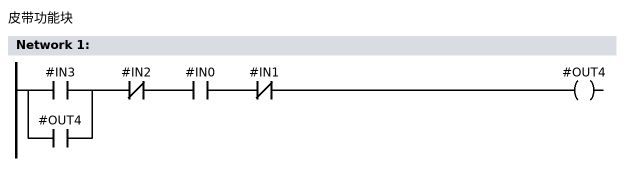
   RUNG wire#powerrail
      Contact( #IN3 )
      wire#w1
      I_Contact( #IN2 )
      Contact( #IN0 )
      I_Contact( #IN1 )
      Coil( #OUT4 )
   END_RUNG
   RUNG wire#powerrail
      Contact( #OUT4 )
   END_RUNG wire#w1
   // the same network as SCL:
   #OUT4 := (#IN3 OR #OUT4) AND NOT #IN2 AND #IN0 AND NOT #IN1;
END_REGION
END_FUNCTION

FUNCTION "脉冲累计功能块" : Void   // FC116, LAD
{ S7_Optimized_Access := 'FALSE' }
VERSION : 0.1
   VAR_INPUT
      IN0 : Bool;
      IN1 : Bool;
   END_VAR
   VAR_OUTPUT
      OUT2 : Real;
   END_VAR
   VAR_TEMP
      TEMP3 : Bool;
      TEMP4 : Real;
      TEMP5 : Real;
      TEMP6 : Real;
   END_VAR
   VAR_TEMP   // added for the SCL form of the ladder/FBD networks
      _w1 : Bool;
   END_VAR
BEGIN

REGION Network 2
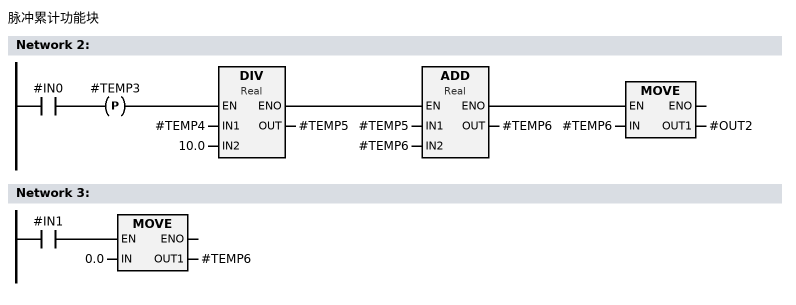
   RUNG wire#powerrail
      Contact( #IN0 )
      P_Trig( #TEMP3 )
      { S7_Templates := "SrcType := Real"; S7_GenerateENO := "TRUE" } Div(in1 := #TEMP4, in2 := 10.0, out => #TEMP5)
      { S7_Templates := "SrcType := Real"; S7_GenerateENO := "TRUE" } Add(in1 := #TEMP5, in2 := #TEMP6, out => #TEMP6)
      { S7_GenerateENO := "TRUE" } Move(in := #TEMP6, out1 => #OUT2)
   END_RUNG
   // the same network as SCL:
   // ENO of a box is taken as its EN; it also drops when the box reports an error
   #_w1 := #IN0 AND NOT #TEMP3;   // rising edge
   #TEMP3 := #IN0;
   IF #_w1 THEN
       #TEMP5 := #TEMP4 / 10.0;
       #TEMP6 := #TEMP5 + #TEMP6;
       #OUT2 := #TEMP6;
   END_IF;
END_REGION

REGION Network 3
   RUNG wire#powerrail
      Contact( #IN1 )
      { S7_GenerateENO := "TRUE" } Move(in := 0.0, out1 => #TEMP6)
   END_RUNG
   // the same network as SCL:
   IF #IN1 THEN #TEMP6 := 0.0; END_IF;
END_REGION

REGION Network 4 (STL)
         SET;
         SAVE;
END_REGION
END_FUNCTION

ORGANIZATION_BLOCK "Main"   // OB1, LAD, ProgramCycle
{ S7_Optimized_Access := 'FALSE' }
VERSION : 0.1
   VAR_TEMP
      TEMP0 : Byte;
      TEMP1 : Byte;
      TEMP2 : Byte;
      TEMP3 : Byte;
      TEMP4 : Byte;
      TEMP5 : Byte;
      TEMP6 : Int;
      TEMP7 : Int;
      TEMP8 : Int;
      TEMP9 : Date_And_Time;
   END_VAR
BEGIN

REGION Network 1
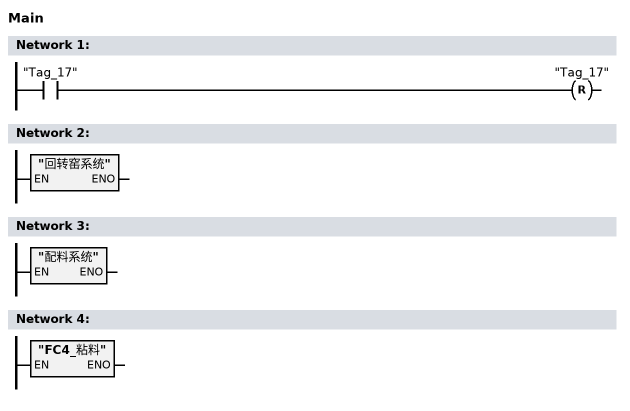
   RUNG wire#powerrail
      Contact( "Tag_17" )
      R_Coil( "Tag_17" )
   END_RUNG
   // the same network as SCL:
   IF "Tag_17" THEN "Tag_17" := FALSE; END_IF;
END_REGION

REGION Network 2
   RUNG wire#powerrail
      "回转窑系统"()
   END_RUNG
   // the same network as SCL:
   "回转窑系统"();
END_REGION

REGION Network 3
   RUNG wire#powerrail
      "配料系统"()
   END_RUNG
   // the same network as SCL:
   "配料系统"();
END_REGION

REGION Network 4
   RUNG wire#powerrail
      "FC4_粘料"()
   END_RUNG
   // the same network as SCL:
   "FC4_粘料"();
END_REGION
END_ORGANIZATION_BLOCK

ORGANIZATION_BLOCK "Cyclic interrupt"   // OB30, LAD, CyclicInterrupt
{ S7_Optimized_Access := 'TRUE' }
VERSION : 0.1
   VAR_INPUT
      Initial_Call : Bool;   // Initial call of this OB
      Event_Count : Int;   // Events discarded
   END_VAR
   VAR_TEMP   // added for the SCL form of the ladder/FBD networks
      _w1 : Bool;
      _w2 : Bool;
   END_VAR
BEGIN

REGION Network 1
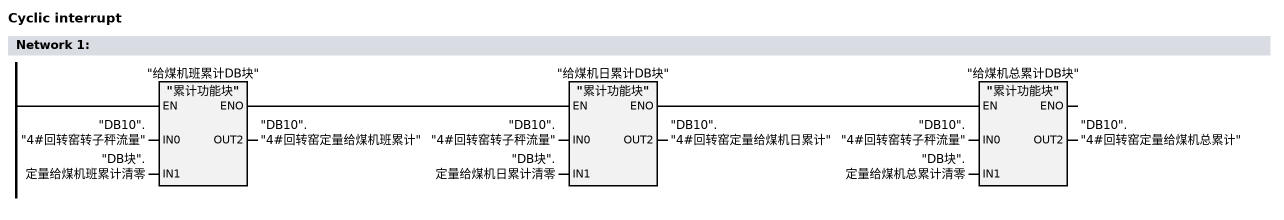
   RUNG wire#powerrail
      "给煤机班累计DB块"(IN0 := "DB10"."4#回转窑转子秤流量", IN1 := "DB块".定量给煤机班累计清零, OUT2 => "DB10"."4#回转窑定量给煤机班累计")
      "给煤机日累计DB块"(IN0 := "DB10"."4#回转窑转子秤流量", IN1 := "DB块".定量给煤机日累计清零, OUT2 => "DB10"."4#回转窑定量给煤机日累计")
      "给煤机总累计DB块"(IN0 := "DB10"."4#回转窑转子秤流量", IN1 := "DB块".定量给煤机总累计清零, OUT2 => "DB10"."4#回转窑定量给煤机总累计")
   END_RUNG
   // the same network as SCL:
   "给煤机班累计DB块"(IN0 := "DB10"."4#回转窑转子秤流量", IN1 := "DB块".定量给煤机班累计清零, OUT2 => "DB10"."4#回转窑定量给煤机班累计", ENO => #_w1);   // "累计功能块"
   "给煤机日累计DB块"(EN := #_w1,   // "累计功能块"
               IN0 := "DB10"."4#回转窑转子秤流量",
               IN1 := "DB块".定量给煤机日累计清零,
               OUT2 => "DB10"."4#回转窑定量给煤机日累计",
               ENO => #_w2);
   IF #_w2 THEN
       "给煤机总累计DB块"(IN0 := "DB10"."4#回转窑转子秤流量", IN1 := "DB块".定量给煤机总累计清零, OUT2 => "DB10"."4#回转窑定量给煤机总累计");   // "累计功能块"
   END_IF;
END_REGION
END_ORGANIZATION_BLOCK

// ===== PLC "1#LM"  CPU 1511-1 PN =====

VAR_GLOBAL   // PLC tag table "默认变量表"
   "送煤皮带备妥" AT %I0.0 : Bool;
   "送煤皮带运行" AT %I0.1 : Bool;
   "送煤皮带故障" AT %I0.2 : Bool;
   "除铁器备妥" AT %I0.3 : Bool;
   "除铁器运行" AT %I0.4 : Bool;
   "除铁器故障" AT %I0.5 : Bool;
   "定量给煤机备妥" AT %I0.6 : Bool;
   "定量给煤机运行" AT %I0.7 : Bool;
   "定量给煤机故障" AT %I1.0 : Bool;
   "煤粉收尘器备妥" AT %I1.1 : Bool;
   "煤粉收尘器运行" AT %I1.2 : Bool;
   "煤粉收尘器故障" AT %I1.3 : Bool;
   "立磨尾排风机远程" AT %I1.4 : Bool;
   "立磨尾排风机运行" AT %I1.5 : Bool;
   "立磨尾排风机故障" AT %I1.6 : Bool;
   "立磨尾排风机待机" AT %I1.7 : Bool;
   "立磨尾排高压柜远程" AT %I2.0 : Bool;
   "立磨尾排高压柜合闸" AT %I2.1 : Bool;
   "立磨尾排高压柜分闸" AT %I2.2 : Bool;
   "定量给煤机断料信号" AT %I2.3 : Bool;
   "定量给煤机左跑偏信号" AT %I2.4 : Bool;
   "定量给煤机右跑偏信号" AT %I2.5 : Bool;
   "给煤机断链信号" AT %I2.6 : Bool;
   "立磨给煤机累计脉冲" AT %I2.7 : Bool;
   "定量给料机远程" AT %I3.0 : Bool;
   "1#铰刀运行" AT %I3.1 : Bool;
   "2#铰刀运行" AT %I3.2 : Bool;
   "1#分割轮运行" AT %I3.3 : Bool;
   "2#分割轮运行" AT %I3.4 : Bool;
   "3#分割轮运行" AT %I3.5 : Bool;
   "4#分割轮运行" AT %I3.6 : Bool;
   "5#分割轮运行" AT %I3.7 : Bool;
   "立磨主机高压柜远程" AT %I4.0 : Bool;
   "立磨主机高压柜合闸" AT %I4.1 : Bool;
   "立磨主机高压柜分闸" AT %I4.2 : Bool;
   "立磨主机运行" AT %I4.3 : Bool;
   "立磨主机故障" AT %I4.4 : Bool;
   "允许主机启动" AT %I4.5 : Bool;
   "停主机" AT %I4.6 : Bool;
   "6#分割轮运行" AT %I5.0 : Bool;
   "7#分割轮运行" AT %I5.1 : Bool;
   "8#分割轮运行" AT %I5.2 : Bool;
   "9#分割轮运行" AT %I5.3 : Bool;
   "10#分割轮运行" AT %I5.4 : Bool;
   "1#灰管压力" AT %IW112 : Word;
   "2#灰管压力" AT %IW114 : Word;
   "Tag_76" AT %IW116 : Word;
   "Tag_78" AT %IW118 : Word;
   "1#母管压力USELESS" AT %IW212 : Word;
   "1#灰管压力UEELESS" AT %IW214 : Word;
   "2#母管压力USELESS" AT %IW216 : Word;
   "2#灰管压力USELESS" AT %IW218 : Word;
   "立磨尾排风机水平震动1" AT %IW256 : Int;
   "立磨尾排风机水平震动2" AT %IW258 : Int;
   "立磨尾排风机垂直震动1" AT %IW260 : Int;
   "立磨尾排风机垂直震动2" AT %IW262 : Int;
   "立磨尾排风机入口压力1" AT %IW264 : Int;
   "立磨尾排风机入口压力2" AT %IW266 : Int;
   "立磨尾排风机出口压力1" AT %IW268 : Int;
   "尾排风机入口执行器反馈" AT %IW270 : Int;
   "立磨1#煤粉仓负压" AT %IW272 : Int;
   "立磨2#煤粉仓负压" AT %IW274 : Int;
   "立磨热风管道负压" AT %IW276 : Int;
   "立磨主电机运行电流" AT %IW278 : Int;
   "立磨给煤机流量" AT %IW280 : Int;
   "立磨出口压力1" AT %IW282 : Int;
   "立磨出口压力2" AT %IW284 : Int;
   "立磨尾排风机运行转速" AT %IW288 : Int;
   "立磨尾排风机运行电流" AT %IW290 : Int;
   "立磨尾排风机出口温度1" AT %IW292 : Int;
   "立磨尾排风机入口温度1" AT %IW296 : Int;
   "立磨尾排风机入口温度2" AT %IW298 : Int;
   "立磨入磨口温度" AT %IW300 : Int;
   "1#煤粉仓1#温度" AT %ID304 : DWord;
   "1#煤粉仓2#温度" AT %ID308 : DWord;
   "1#煤粉仓3#温度" AT %ID312 : DWord;
   "1#煤粉仓4#温度" AT %ID316 : DWord;
   "1#煤粉仓5#温度" AT %ID320 : DWord;
   "1#煤粉仓6#温度" AT %ID324 : DWord;
   "2#煤粉仓1#温度" AT %ID328 : DWord;
   "2#煤粉仓2#温度" AT %ID332 : DWord;
   "2#煤粉仓3#温度" AT %ID336 : DWord;
   "2#煤粉仓4#温度" AT %ID340 : DWord;
   "2#煤粉仓5#温度" AT %ID344 : DWord;
   "2#煤粉仓6#温度" AT %ID348 : DWord;
   "电机绕组U相温度" AT %ID352 : DWord;
   "电机绕组V相温度" AT %ID356 : DWord;
   "电机绕组W相温度" AT %ID360 : DWord;
   "尾排电机前轴温度" AT %ID364 : DWord;
   "尾排电机后轴温度" AT %ID368 : DWord;
   "尾排风机前轴温度" AT %ID372 : DWord;
   "尾排风机后轴温度" AT %ID376 : DWord;
   "立磨机出口温度1" AT %ID380 : DWord;
   "立磨机出口温度2" AT %ID384 : DWord;
   "Tag_101" AT %ID388 : DWord;
   "Tag_102" AT %ID392 : DWord;
   "Tag_103" AT %ID396 : DWord;
   "送煤皮带驱动" AT %Q0.0 : Bool;
   "除铁器驱动" AT %Q0.1 : Bool;
   "定量给煤机驱动" AT %Q0.2 : Bool;
   "煤粉收尘器驱动" AT %Q0.3 : Bool;
   "立磨尾排风机停止" AT %Q0.4 : Bool;
   "立磨尾排高压柜合闸驱动" AT %Q0.5 : Bool;
   "立磨尾排风机高压柜分闸" AT %Q0.6 : Bool;
   "立磨尾排风机驱动" AT %Q0.7 : Bool;
   "立磨主机高压柜合闸驱动" AT %Q1.0 : Bool;
   "立磨主机高压柜分闸驱动" AT %Q1.1 : Bool;
   "Tag_107" AT %QB4 : Byte;
   "1#仓泵手/自动" AT %Q100.0 : Bool;
   "1#仓泵自动启动" AT %Q100.1 : Bool;
   "1#仓泵自动停止" AT %Q100.2 : Bool;
   "2#仓泵手/自动" AT %Q100.3 : Bool;
   "2#仓泵自动启动" AT %Q100.4 : Bool;
   "2#仓泵自动停止" AT %Q100.5 : Bool;
   "1#排气阀手动开" AT %Q101.0 : Bool;
   "1#排气阀手动关" AT %Q101.1 : Bool;
   "1#进料阀手动开" AT %Q101.2 : Bool;
   "1#进料阀手动关" AT %Q101.3 : Bool;
   "1#出料阀手动开" AT %Q101.4 : Bool;
   "1#出料阀手动关" AT %Q101.5 : Bool;
   "1#进气阀手动开" AT %Q101.6 : Bool;
   "1#进气阀手动关" AT %Q101.7 : Bool;
   "1#助吹阀手动开" AT %Q102.0 : Bool;
   "1#助吹阀手动关" AT %Q102.1 : Bool;
   "1#排堵阀手动开" AT %Q102.2 : Bool;
   "1#排堵阀手动关" AT %Q102.3 : Bool;
   "2#排气阀手动开" AT %Q102.4 : Bool;
   "2#排气阀手动关" AT %Q102.5 : Bool;
   "2#进料阀手动开" AT %Q102.6 : Bool;
   "2#进料阀手动关" AT %Q102.7 : Bool;
   "2#出料阀手动开" AT %Q103.0 : Bool;
   "2#出料阀手动关" AT %Q103.1 : Bool;
   "2#进气阀手动开" AT %Q103.2 : Bool;
   "2#进气阀手动关" AT %Q103.3 : Bool;
   "2#助吹阀手动开" AT %Q103.4 : Bool;
   "2#助吹阀手动关" AT %Q103.5 : Bool;
   "2#排堵阀手动开" AT %Q103.6 : Bool;
   "2#排堵阀手动关" AT %Q103.7 : Bool;
   "1#切1#切换阀手动开" AT %Q104.0 : Bool;
   "1#切1#切换阀手动关" AT %Q104.1 : Bool;
   "1#切2#切换阀手动开" AT %Q104.2 : Bool;
   "1#切2#切换阀手动关" AT %Q104.3 : Bool;
   "1#切3#切换阀手动开" AT %Q104.4 : Bool;
   "1#切3#切换阀手动关" AT %Q104.5 : Bool;
   "1#切4#切换阀手动开" AT %Q104.6 : Bool;
   "1#切4#切换阀手动关" AT %Q104.7 : Bool;
   "1#切5#切换阀手动开" AT %Q105.0 : Bool;
   "1#切5#切换阀手动关" AT %Q105.1 : Bool;
   "2#切1#切换阀手动开" AT %Q105.2 : Bool;
   "2#切1#切换阀手动关" AT %Q105.3 : Bool;
   "2#切2#切换阀手动开" AT %Q105.4 : Bool;
   "1#母管压力下限" AT %QW108 : Word;
   "1#灰管压力下限" AT %QW110 : Word;
   "1#灰管压力上限" AT %QW112 : Word;
   "1#进料时间" AT %QW114 : Word;
   "1#吹扫时间" AT %QW116 : Word;
   "2#母管压力下限" AT %QW118 : Word;
   "2#灰管压力下限" AT %QW120 : Word;
   "2#灰管压力上限" AT %QW122 : Word;
   "2#进料时间" AT %QW124 : Word;
   "立磨给煤机流量给定" AT %QW256 : Int;
   "立磨尾排风机转速给定" AT %QW258 : Int;
   "尾排风机入口执行器给定" AT %QW260 : Int;
   "Tag_5" AT %M2.0 : Bool;
   "Tag_11" AT %M2.3 : Bool;
   "Tag_19" AT %M2.5 : Bool;
   "Tag_1" AT %MW4 : Word;
   "Tag_8" AT %MW10 : Word;
   "Tag_6" AT %MW12 : Word;
   "Tag_21" AT %MW14 : Word;
   "Tag_16" AT %MW16 : Word;
   "锁风定量给煤机流量累计清零" AT %M30.1 : Bool;
   "Tag_13" AT %MW100 : Word;
   "Tag_12" AT %M300.0 : Bool;
   "Tag_20" AT %M300.1 : Bool;
   "Tag_9" AT %M400.0 : Bool;
   "Tag_17" AT %M400.1 : Bool;
   "1#仓泵进料时间" AT %MW506 : Word;
   "1#仓泵吹扫时间" AT %MW508 : Word;
   "1#母管下限" AT %MW510 : Word;
   "1#灰管上限" AT %MW512 : Word;
   "1#灰管下限" AT %MW514 : Word;
   "2#仓泵进料时间" AT %MW516 : Word;
   "2#仓泵吹扫时间" AT %MW518 : Word;
   "2#母管下限" AT %MW520 : Word;
   "2#灰管上限" AT %MW522 : Word;
   "2#灰管下限" AT %MW524 : Word;
   "1#母管压力信号" AT %MW526 : Word;
   "1#灰管压力信号" AT %MW528 : Word;
   "2#母管压力信号" AT %MW530 : Word;
   "2#灰管压力信号" AT %MW532 : Word;
   "1#仓泵手自动标示" AT %M600.1 : Bool;
   "2#仓泵手自动标示" AT %M600.2 : Bool;
   "Tag_3" AT %T100 : Timer;
   "Tag_4" AT %T101 : Timer;
   "Tag_10" AT %C1 : Counter;
   "Tag_18" AT %C2 : Counter;
   "I4_7" AT %I4.7 : Bool;
   "I5_5" AT %I5.5 : Bool;
   "I5_6" AT %I5.6 : Bool;
   "I5_7" AT %I5.7 : Bool;
   "1#板式给煤机-褐煤备妥" AT %I6.0 : Bool;
   "1#板式给煤机-褐煤运行" AT %I6.1 : Bool;
   "1#板式给煤机-褐煤故障" AT %I6.2 : Bool;
   "2#板式给煤机-烟煤备妥" AT %I6.3 : Bool;
   "2#板式给煤机-烟煤运行" AT %I6.4 : Bool;
   "2#板式给煤机-烟煤故障" AT %I6.5 : Bool;
   "I6_6" AT %I6.6 : Bool;
   "I6_7" AT %I6.7 : Bool;
   "I7_0" AT %I7.0 : Bool;
   "I7_1" AT %I7.1 : Bool;
   "I7_2" AT %I7.2 : Bool;
   "I7_3" AT %I7.3 : Bool;
   "I7_4" AT %I7.4 : Bool;
   "I7_5" AT %I7.5 : Bool;
   "I7_6" AT %I7.6 : Bool;
   "I7_7" AT %I7.7 : Bool;
   "I8_0" AT %I8.0 : Bool;
   "I8_1" AT %I8.1 : Bool;
   "I8_2" AT %I8.2 : Bool;
   "I8_3" AT %I8.3 : Bool;
   "I8_4" AT %I8.4 : Bool;
   "I8_5" AT %I8.5 : Bool;
   "I8_6" AT %I8.6 : Bool;
   "I8_7" AT %I8.7 : Bool;
   "I9_0" AT %I9.0 : Bool;
   "I9_1" AT %I9.1 : Bool;
   "I9_2" AT %I9.2 : Bool;
   "I9_3" AT %I9.3 : Bool;
   "I9_4" AT %I9.4 : Bool;
   "I9_5" AT %I9.5 : Bool;
   "I9_6" AT %I9.6 : Bool;
   "I9_7" AT %I9.7 : Bool;
   "I10_0" AT %I10.0 : Bool;
   "I10_1" AT %I10.1 : Bool;
   "I10_2" AT %I10.2 : Bool;
   "I10_3" AT %I10.3 : Bool;
   "I10_4" AT %I10.4 : Bool;
   "I10_5" AT %I10.5 : Bool;
   "I10_6" AT %I10.6 : Bool;
   "I10_7" AT %I10.7 : Bool;
   "I11_0" AT %I11.0 : Bool;
   "I11_1" AT %I11.1 : Bool;
   "I11_2" AT %I11.2 : Bool;
   "I11_3" AT %I11.3 : Bool;
   "I11_4" AT %I11.4 : Bool;
   "I11_5" AT %I11.5 : Bool;
   "I11_6" AT %I11.6 : Bool;
   "I11_7" AT %I11.7 : Bool;
   "1#板式给煤机-褐煤启停" AT %Q1.2 : Bool;
   "2#板式给煤机-烟煤启停" AT %Q1.3 : Bool;
   "立磨现场皮带报警器" AT %Q1.4 : Bool;
   "立磨中控报警器" AT %Q1.5 : Bool;
   "Q1_6" AT %Q1.6 : Bool;
   "Q1_7" AT %Q1.7 : Bool;
   "Q2_0" AT %Q2.0 : Bool;
   "Q2_1" AT %Q2.1 : Bool;
   "Q2_2" AT %Q2.2 : Bool;
   "Q2_3" AT %Q2.3 : Bool;
   "Q2_4" AT %Q2.4 : Bool;
   "Q2_5" AT %Q2.5 : Bool;
   "Q2_6" AT %Q2.6 : Bool;
   "Q2_7" AT %Q2.7 : Bool;
   "Q3_0" AT %Q3.0 : Bool;
   "Q3_1" AT %Q3.1 : Bool;
   "Q3_2" AT %Q3.2 : Bool;
   "Q3_3" AT %Q3.3 : Bool;
   "Q3_4" AT %Q3.4 : Bool;
   "Q3_5" AT %Q3.5 : Bool;
   "Q3_6" AT %Q3.6 : Bool;
   "Q3_7" AT %Q3.7 : Bool;
   "1#板式给煤机-褐煤流量反馈" AT %IW286 : Int;
   "2#板式给煤机-烟煤流量反馈" AT %IW294 : Int;
   "PIW302" AT %IW302 : Int;
   "1#板式给煤机-褐煤流量给定" AT %QW262 : Int;
   "2#板式给煤机-烟煤流量给定" AT %QW264 : Int;
   "PQW266" AT %QW266 : Int;
   "PQW268" AT %QW268 : Int;
   "PQW270" AT %QW270 : Int;
   "立磨煤粉仓称重" AT %ID400 : Real;
   "立磨1#煤粉仓称重" AT %ID408 : Real;
   "立磨2#煤粉仓称重" AT %ID416 : Real;
   "1#立磨板式给料流量累计清零" AT %M30.2 : Bool;
   "2#立磨板式给料流量累计清零" AT %M30.3 : Bool;
   "Tag_2" AT %M30.7 : Bool;
   "Tag_80" AT %M80.0 : Bool;
   "Tag_81" AT %M81.0 : Bool;
   "Tag_82" AT %M80.1 : Bool;
   "Tag_83" AT %M80.2 : Bool;
   "Tag_84" AT %M80.3 : Bool;
   "Tag_85" AT %M81.1 : Bool;
   "Tag_86" AT %T102 : Timer;
   "Clock_Byte" AT %MB0 : Byte;
   "Clock_10Hz" AT %M0.0 : Bool;
   "Clock_5Hz" AT %M0.1 : Bool;
   "Clock_2.5Hz" AT %M0.2 : Bool;
   "Clock_2Hz" AT %M0.3 : Bool;
   "Clock_1.25Hz" AT %M0.4 : Bool;
   "Clock_1Hz" AT %M0.5 : Bool;
   "Clock_0.625Hz" AT %M0.6 : Bool;
   "Clock_0.5Hz" AT %M0.7 : Bool;
   "System_Byte" AT %MB1 : Byte;
   "FirstScan" AT %M1.0 : Bool;
   "DiagStatusUpdate" AT %M1.1 : Bool;
   "AlwaysTRUE" AT %M1.2 : Bool;
   "AlwaysFALSE" AT %M1.3 : Bool;
   "2#切2#切换阀手动关" AT %Q105.5 : Bool;
   "3#切1#切换阀手动开" AT %Q105.6 : Bool;
   "3#切1#切换阀手动关" AT %Q105.7 : Bool;
   "3#切2#切换阀手动开" AT %Q106.0 : Bool;
   "3#切2#切换阀手动关" AT %Q106.1 : Bool;
   "4#切1#切换阀手动开" AT %Q106.2 : Bool;
   "4#切1#切换阀手动关" AT %Q106.3 : Bool;
   "4#切2#切换阀手动开" AT %Q106.4 : Bool;
   "4#切2#切换阀手动关" AT %Q106.5 : Bool;
   "4#切3#切换阀手动开" AT %Q106.6 : Bool;
   "4#切3#切换阀手动关" AT %Q106.7 : Bool;
   "4#切4#切换阀手动开" AT %Q107.0 : Bool;
   "4#切4#切换阀手动关" AT %Q107.1 : Bool;
   "Tag_20(1)" AT %Q107.2 : Bool;
   "Tag_21(1)" AT %Q107.3 : Bool;
   "Tag_22" AT %Q107.4 : Bool;
   "Tag_23" AT %Q107.5 : Bool;
   "Tag_24" AT %Q107.6 : Bool;
   "Tag_25" AT %Q107.7 : Bool;
   "2#吹扫时间" AT %QW126 : Word;
   "1#排气阀关到位" AT %I100.0 : Bool;
   "1#排气阀开到位" AT %I100.1 : Bool;
   "1#进料阀关到位" AT %I100.2 : Bool;
   "1#进料阀开到位" AT %I100.3 : Bool;
   "1#出料阀关到位" AT %I100.4 : Bool;
   "1#出料阀开到位" AT %I100.5 : Bool;
   "1#进气阀关到位" AT %I100.6 : Bool;
   "1#进气阀开到位" AT %I100.7 : Bool;
   "1#助吹阀关到位" AT %I101.0 : Bool;
   "1#助吹阀开到位" AT %I101.1 : Bool;
   "1#排堵阀关到位" AT %I101.2 : Bool;
   "1#排堵阀开到位" AT %I101.3 : Bool;
   "1#料位信号" AT %I101.4 : Bool;
   "1#现场箱远程" AT %I101.5 : Bool;
   "2#排气阀关到位" AT %I101.6 : Bool;
   "2#排气阀开到位" AT %I101.7 : Bool;
   "2#进料阀关到位" AT %I102.0 : Bool;
   "2#进料阀开到位" AT %I102.1 : Bool;
   "2#出料阀关到位" AT %I102.2 : Bool;
   "2#出料阀开到位" AT %I102.3 : Bool;
   "2#进气阀关到位" AT %I102.4 : Bool;
   "2#进气阀开到位" AT %I102.5 : Bool;
   "2#助吹阀关到位" AT %I102.6 : Bool;
   "2#助吹阀开到位" AT %I102.7 : Bool;
   "2#排堵阀关到位" AT %I103.0 : Bool;
   "2#排堵阀开到位" AT %I103.1 : Bool;
   "2#料位信号" AT %I103.2 : Bool;
   "2#现场箱远程" AT %I103.3 : Bool;
   "1#切1#切换阀关到位" AT %I103.4 : Bool;
   "1#切1#切换阀开到位" AT %I103.5 : Bool;
   "1#切2#切换阀关到位" AT %I103.6 : Bool;
   "1#切2#切换阀开到位" AT %I103.7 : Bool;
   "1#切3#切换阀关到位" AT %I104.0 : Bool;
   "1#切3#切换阀开到位" AT %I104.1 : Bool;
   "1#切4#切换阀关到位" AT %I104.2 : Bool;
   "1#切4#切换阀开到位" AT %I104.3 : Bool;
   "1#切5#切换阀关到位" AT %I104.4 : Bool;
   "1#切5#切换阀开到位" AT %I104.5 : Bool;
   "1#切远程信号" AT %I104.6 : Bool;
   "2#切1#切换阀关到位" AT %I104.7 : Bool;
   "2#切1#切换阀开到位" AT %I105.0 : Bool;
   "2#切2#切换阀关到位" AT %I105.1 : Bool;
   "2#切2#切换阀开到位" AT %I105.2 : Bool;
   "2#切远程信号" AT %I105.3 : Bool;
   "3#切1#切换阀关到位" AT %I105.4 : Bool;
   "3#切1#切换阀开到位" AT %I105.5 : Bool;
   "3#切2#切换阀关到位" AT %I105.6 : Bool;
   "3#切2#切换阀开到位" AT %I105.7 : Bool;
   "3#切远程信号" AT %I106.0 : Bool;
   "4#切1#切换阀关到位" AT %I106.1 : Bool;
   "4#切1#切换阀开到位" AT %I106.2 : Bool;
   "4#切2#切换阀关到位" AT %I106.3 : Bool;
   "4#切2#切换阀开到位" AT %I106.4 : Bool;
   "4#切3#切换阀关到位" AT %I106.5 : Bool;
   "4#切3#切换阀开到位" AT %I106.6 : Bool;
   "4#切4#切换阀关到位" AT %I106.7 : Bool;
   "4#切4#切换阀开到位" AT %I107.0 : Bool;
   "4#切远程信号" AT %I107.1 : Bool;
   "1#中控备妥" AT %I107.2 : Bool;
   "1#运行" AT %I107.3 : Bool;
   "1#母管压力低" AT %I107.4 : Bool;
   "1#灰管压力高" AT %I107.5 : Bool;
   "2#中控备妥" AT %I107.6 : Bool;
   "2#运行" AT %I107.7 : Bool;
   "2#母管压力低" AT %I108.0 : Bool;
   "2#灰管压力高" AT %I108.1 : Bool;
   "Tag_7" AT %MW200 : Word;
   "Tag_14" AT %MW202 : Word;
   "Tag_15" AT %M200.0 : Bool;
   "Tag_26" AT %M200.1 : Bool;
   "Tag_27" AT %Q4.0 : Bool;
   "Tag_28" AT %M2.1 : Bool;
   "Tag_29" AT %MW82 : Word;
   "Tag_30" AT %C3 : Counter;
   "Tag_31" AT %C4 : Counter;
   "母管压力" AT %IW110 : Word;
   "Tag_32" AT %M10.0 : Bool;
   "Tag_33" AT %MD40 : Real;
   "Tag_34" AT %MD44 : Real;
   "Tag_35" AT %MD48 : Real;
   "Tag_36" AT %M60.0 : Bool;
   "HMI_ALARM_RST" AT %M10.1 : Bool;
   "Tag_38" AT %M10.2 : Bool;
END_VAR

DATA_BLOCK "qud"   // DB1
{ S7_Optimized_Access := 'FALSE' }
VERSION : 0.1
   VAR
      STAT0 : Bool;
      STAT1 : Bool;
      STAT2 : Bool;
      STAT3 : Bool;
      STAT4 : Bool;
      STAT5 : Bool;
      STAT6 : Bool;
      STAT7 : Bool;
      STAT8 : Bool;
      STAT9 : Bool;
      STAT10 : Bool;
      STAT11 : Bool;
      STAT12 : Bool;
      STAT13 : Bool;
      STAT14 : Bool;
      STAT15 : Bool;
      "1#立磨板式给料机启动" : Bool;
      "1#立磨板式给料机停止" : Bool;
      "2#立磨板式给料机启动" : Bool;
      "2#立磨板式给料机停止" : Bool;
      STAT20 : Bool;
      STAT21 : Bool;
      STAT22 : Bool;
      STAT23 : Bool;
   END_VAR
BEGIN
END_DATA_BLOCK

DATA_BLOCK "MNL"   // DB2
{ S7_Optimized_Access := 'FALSE' }
VERSION : 0.1
   VAR
      锁风定量给煤机 : Real := 44.0;
      锁风定量给煤机流量反馈 : Real;
      立磨尾排水平振动1 : Real;
      立磨尾排水平振动2 : Real;
      立磨尾排风机垂直振动1 : Real;
      立磨尾排风机垂直振动2 : Real;
      立磨尾排风机出口压力1 : Real;
      立磨尾排风机出口压力2 : Real;
      STAT8 : Real := 56.07639;
      立磨尾排风机出口温度2 : Real;
      STAT10 : Real := 47.39583;
      STAT11 : Real := 46.52778;
      立磨尾排风机入口压力1 : Real := -2147.512;
      立磨尾排风机入口压力2 : Real := -2461.689;
      "立磨1#煤粉仓负压" : Real := -300.0;
      "立磨2#煤粉仓负压" : Real := -272.9167;
      立磨热风管道负压 : Real := -562.5;
      立磨煤粉仓称重 : Real := 101.51;
      "立磨1#煤粉仓称重" : Real := 8.44;
      "立磨2#煤粉仓称重" : Real := 13.24;
      尾排风机运行频率 : Real := 744.2824;
      尾排风机运行电流 : Real := 41.25;
      主电机运行电流 : Real;
      立磨尾排风机转速给定 : Real := 500.0;
      锁风定量给煤机流量累计 : Real := 30006.97;
      "1#煤粉仓1#温度" : Real := 37.0;
      "1#煤粉仓2#温度" : Real := 36.0;
      "1#煤粉仓3#温度" : Real := 37.0;
      "1#煤粉仓4#温度" : Real := 36.0;
      "1#煤粉仓5#温度" : Real := 36.0;
      "1#煤粉仓6#温度" : Real := 37.0;
      "2#煤粉仓1#温度" : Real := 37.0;
      "2#煤粉仓2#温度" : Real := 36.0;
      "2#煤粉仓3#温度" : Real := 37.0;
      "2#煤粉仓4#温度" : Real := 37.0;
      "2#煤粉仓5#温度" : Real := 37.0;
      "2#煤粉仓6#温度" : Real := 37.0;
      电机绕组U相温度 : Real := 59.0;
      电机绕组V相温度 : Real := 57.0;
      电机绕组W相温度 : Real := 59.0;
      尾排电机前轴温度 : Real := 34.0;
      尾排电机后轴温度 : Real := 40.0;
      尾排风机前轴温度 : Real := 144.8206;
      尾排风机后轴温度 : Real;
      立磨机出口温度1 : Real;
      立磨机出口温度2 : Real := 43.0;
      STAT46 : Real := 46.0;
      STAT47 : Real := 62.0;
      STAT48 : Real := 58.0;
      立磨尾排风机出口温度1 : Real := -1753.472;
      立磨尾排风机入口温度1 : Real := -1707.176;
      立磨尾排风机入口温度2 : Real;
      尾排风机执行器开度给定 : Real;
      尾排风机执行器开度反馈 : Real;
      立磨机出口压力1 : Real;
      立磨机出口压力2 : Real;
      立磨主电机入磨口温度 : Real;
      "1#立磨板式给料反馈" : Real;
      "2#立磨板式给料反馈" : Real;
      "1#立磨板式给料给定" : Real;
      "2#立磨板式给料给定" : Real;
      "1#立磨板式给料累计" : Real;
      "2#立磨板式给料累计" : Real;
      STAT63 : Real;
      STAT64 : Real;
      STAT65 : Real;
   END_VAR
BEGIN
END_DATA_BLOCK

DATA_BLOCK "TIMEDB"   // DB3
{ S7_Optimized_Access := 'TRUE' }
VERSION : 0.1
   VAR
      T1 : IEC_TIMER;
      T2 : IEC_TIMER;
      T3 : IEC_TIMER;
      T4 : IEC_TIMER;
      T5 : IEC_TIMER;
      T6 : IEC_TIMER;
      T7 : IEC_TIMER;
      T8 : IEC_TIMER;
      T9 : IEC_TIMER;
      T10 : IEC_TIMER;
      T11 : IEC_TIMER;
      T12 : IEC_TIMER;
      T13 : IEC_TIMER;
      T14 : IEC_TIMER;
      T15 : IEC_TIMER;
      T16 : IEC_TIMER;
      T17 : IEC_TIMER;
      T18 : IEC_TIMER;
      T19 : IEC_TIMER;
      T20 : IEC_TIMER;
      T21 : IEC_TIMER;
      T22 : IEC_TIMER;
      T23 : IEC_TIMER;
      T24 : IEC_TIMER;
      T25 : IEC_TIMER;
      T26 : IEC_TIMER;
      T27 : IEC_TIMER;
      T28 : IEC_TIMER;
      T29 : IEC_TIMER;
      T30 : IEC_TIMER;
      T31 : IEC_TIMER;
      T32 : IEC_TIMER;
      T33 : IEC_TIMER;
      T34 : IEC_TIMER;
      T35 : IEC_TIMER;
      T36 : IEC_TIMER;
      T37 : IEC_TIMER;
      T38 : IEC_TIMER;
      T39 : IEC_TIMER;
      T40 : IEC_TIMER;
      T41 : IEC_TIMER;
      T42 : IEC_TIMER;
      T43 : IEC_TIMER;
      T44 : IEC_TIMER;
      T45 : IEC_TIMER;
      T46 : IEC_TIMER;
      T47 : IEC_TIMER;
      T48 : IEC_TIMER;
      T49 : IEC_TIMER;
      T50 : IEC_TIMER;
      T51 : IEC_TIMER;
      T52 : IEC_TIMER;
      T53 : IEC_TIMER;
      T54 : IEC_TIMER;
      T55 : IEC_TIMER;
      T56 : IEC_TIMER;
      T57 : IEC_TIMER;
      T58 : IEC_TIMER;
      T59 : IEC_TIMER;
      T60 : IEC_TIMER;
      T61 : IEC_TIMER;
      T62 : IEC_TIMER;
      T63 : IEC_TIMER;
      T64 : IEC_TIMER;
      T65 : IEC_TIMER;
      T66 : IEC_TIMER;
      T67 : IEC_TIMER;
      T68 : IEC_TIMER;
      T69 : IEC_TIMER;
      T70 : IEC_TIMER;
      T71 : IEC_TIMER;
      T72 : IEC_TIMER;
      T73 : IEC_TIMER;
      T74 : IEC_TIMER;
      T75 : IEC_TIMER;
      T76 : IEC_TIMER;
      T77 : IEC_TIMER;
      T78 : IEC_TIMER;
      T79 : IEC_TIMER;
      T80 : IEC_TIMER;
      T81 : IEC_TIMER;
      T82 : IEC_TIMER;
      T83 : IEC_TIMER;
      T84 : IEC_TIMER;
      T85 : IEC_TIMER;
      T86 : IEC_TIMER;
      T87 : IEC_TIMER;
      T88 : IEC_TIMER;
      T89 : IEC_TIMER;
      T90 : IEC_TIMER;
      T91 : IEC_TIMER;
      T92 : IEC_TIMER;
      T93 : IEC_TIMER;
      T94 : IEC_TIMER;
      T95 : IEC_TIMER;
      T96 : IEC_TIMER;
      T97 : IEC_TIMER;
      T98 : IEC_TIMER;
      T99 : IEC_TIMER;
      T100 : IEC_TIMER;
   END_VAR
BEGIN
END_DATA_BLOCK

DATA_BLOCK "累计功能块_DB_1"   // DB4
{ S7_Optimized_Access := 'FALSE' }
VERSION : 0.1
// stored: InstanceOfName 累计功能块
"累计功能块"
BEGIN
END_DATA_BLOCK

DATA_BLOCK "累计功能块_DB"   // DB5
{ S7_Optimized_Access := 'FALSE' }
VERSION : 0.1
// stored: InstanceOfName 累计功能块
"累计功能块"
BEGIN
END_DATA_BLOCK

DATA_BLOCK "累计功能块_DB_2"   // DB6
{ S7_Optimized_Access := 'FALSE' }
VERSION : 0.1
// stored: InstanceOfName 累计功能块
"累计功能块"
BEGIN
END_DATA_BLOCK

DATA_BLOCK "DB9_P"   // DB9
{ S7_Optimized_Access := 'FALSE' }
VERSION : 0.1
   VAR
      P1 : Bool;
      P2 : Bool;
      P3 : Bool;
      P4 : Bool;
      P5 : Bool;
      P6 : Bool;
      P7 : Bool;
      P8 : Bool;
      P9 : Bool;
      P10 : Bool;
      P11 : Bool;
      P12 : Bool;
      P13 : Bool;
      P14 : Bool;
      P15 : Bool;
      P16 : Bool;
      P17 : Bool;
      P18 : Bool;
      P19 : Bool;
      P20 : Bool;
      P21 : Bool;
      P22 : Bool;
      P23 : Bool;
      P24 : Bool;
      P25 : Bool;
      P26 : Bool;
      P27 : Bool;
      P28 : Bool;
      P29 : Bool;
      P30 : Bool;
      P31 : Bool;
      P32 : Bool;
      P33 : Bool;
      P34 : Bool;
      P35 : Bool;
      P36 : Bool;
      P37 : Bool;
      P38 : Bool;
      P39 : Bool;
      P40 : Bool;
      P41 : Bool;
      P42 : Bool;
      P43 : Bool;
      P44 : Bool;
      P45 : Bool;
      P46 : Bool;
      P47 : Bool;
      P48 : Bool;
      P49 : Bool;
      P50 : Bool;
      P51 : Bool;
      P52 : Bool;
      P53 : Bool;
      P54 : Bool;
      P55 : Bool;
      P56 : Bool;
      P57 : Bool;
      P58 : Bool;
      P59 : Bool;
      P60 : Bool;
      P61 : Bool;
      P62 : Bool;
      P63 : Bool;
      P64 : Bool;
      P65 : Bool;
      P66 : Bool;
      P67 : Bool;
      P68 : Bool;
      P69 : Bool;
      P70 : Bool;
      P71 : Bool;
      P72 : Bool;
      P73 : Bool;
      P74 : Bool;
      P75 : Bool;
      P76 : Bool;
      P77 : Bool;
      P78 : Bool;
      P79 : Bool;
      P80 : Bool;
      P81 : Bool;
      P82 : Bool;
      P83 : Bool;
      P84 : Bool;
      P85 : Bool;
      P86 : Bool;
      P87 : Bool;
      P88 : Bool;
      P89 : Bool;
      P90 : Bool;
      P91 : Bool;
      P92 : Bool;
      P93 : Bool;
   END_VAR
BEGIN
END_DATA_BLOCK

DATA_BLOCK "HMI_IN_BOOL"   // DB10
{ S7_Optimized_Access := 'FALSE' }
VERSION : 0.1
   VAR
      "1#仓泵手/自动" : Bool;
      "1#仓泵自动启动" : Bool;
      "1#仓泵自动停止" : Bool;
      "2#仓泵手/自动" : Bool;
      "2#仓泵自动启动" : Bool;
      "2#仓泵自动停止" : Bool;
      DB10_0_6 : Bool;
      DB10_0_7 : Bool;
      "1#排气阀手动开" : Bool;
      "1#排气阀手动关" : Bool;
      "1#进料阀手动开" : Bool;
      "1#进料阀手动关" : Bool;
      "1#出料阀手动开" : Bool;
      "1#出料阀手动关" : Bool;
      "1#进气阀手动开" : Bool;
      "1#进气阀手动关" : Bool;
      "1#助吹阀手动开" : Bool;
      "1#助吹阀手动关" : Bool;
      "1#排堵阀手动开" : Bool;
      "1#排堵阀手动关" : Bool;
      "2#排气阀手动开" : Bool;
      "2#排气阀手动关" : Bool;
      "2#进料阀手动开" : Bool;
      "2#进料阀手动关" : Bool;
      "2#出料阀手动开" : Bool;
      "2#出料阀手动关" : Bool;
      "2#进气阀手动开" : Bool;
      "2#进气阀手动关" : Bool;
      "2#助吹阀手动开" : Bool;
      "2#助吹阀手动关" : Bool;
      "2#排堵阀手动开" : Bool;
      "2#排堵阀手动关" : Bool;
      "1#切1#切换阀手动开" : Bool;
      "1#切1#切换阀手动关" : Bool;
      "1#切2#切换阀手动开" : Bool;
      "1#切2#切换阀手动关" : Bool;
      "1#切3#切换阀手动开" : Bool;
      "1#切3#切换阀手动关" : Bool;
      "1#切4#切换阀手动开" : Bool;
      "1#切4#切换阀手动关" : Bool;
      "1#切5#切换阀手动开" : Bool;
      "1#切5#切换阀手动关" : Bool;
      "2#切1#切换阀手动开" : Bool;
      "2#切1#切换阀手动关" : Bool;
      "2#切2#切换阀手动开" : Bool;
      "2#切2#切换阀手动关" : Bool;
      "3#切1#切换阀手动开" : Bool;
      "3#切1#切换阀手动关" : Bool;
      "3#切2#切换阀手动开" : Bool;
      "3#切2#切换阀手动关" : Bool;
      "4#切1#切换阀手动开" : Bool;
      "4#切1#切换阀手动关" : Bool;
      "4#切2#切换阀手动开" : Bool;
      "4#切2#切换阀手动关" : Bool;
      "4#切3#切换阀手动开" : Bool;
      "4#切3#切换阀手动关" : Bool;
      "4#切4#切换阀手动开" : Bool;
      "4#切4#切换阀手动关" : Bool;
      DB10_7_2 : Bool;
      DB10_7_3 : Bool;
      DB10_7_4 : Bool;
      DB10_7_5 : Bool;
      DB10_7_6 : Bool;
      DB10_7_7 : Bool;
      DB10_8_0 : Bool;
      DB10_8_1 : Bool;
      DB10_8_2 : Bool;
      DB10_8_3 : Bool;
      DB10_8_4 : Bool;
      DB10_8_5 : Bool;
      DB10_8_6 : Bool;
      DB10_8_7 : Bool;
      DB10_9_0 : Bool;
      DB10_9_1 : Bool;
      DB10_9_2 : Bool;
      DB10_9_3 : Bool;
      DB10_9_4 : Bool;
      DB10_9_5 : Bool;
      DB10_9_6 : Bool;
      DB10_9_7 : Bool;
      DB10_10_0 : Bool;
      DB10_10_1 : Bool;
      DB10_10_2 : Bool;
      DB10_10_3 : Bool;
      DB10_10_4 : Bool;
      DB10_10_5 : Bool;
      DB10_10_6 : Bool;
      DB10_10_7 : Bool;
      DB_10_11_0 : Bool;
      DB_10_11_1 : Bool;
      DB_10_11_2 : Bool;
      DB_10_11_3 : Bool;
      DB_10_11_4 : Bool;
      DB_10_11_5 : Bool;
      DB_10_11_6 : Bool;
      DB_10_11_7 : Bool;
      DB_10_11_8 : Bool;
      DB_10_11_9 : Bool;
      DB_10_11_10 : Bool;
      DB_10_11_11 : Bool;
      DB_10_11_12 : Bool;
      DB_10_11_13 : Bool;
      DB_10_11_14 : Bool;
      DB_10_11_15 : Bool;
      DB_10_11_16 : Bool;
      DB_10_11_17 : Bool;
      DB_10_11_18 : Bool;
      DB_10_11_19 : Bool;
      DB_10_11_20 : Bool;
      DB_10_11_21 : Bool;
      DB_10_11_22 : Bool;
      DB_10_11_23 : Bool;
      DB_10_11_24 : Bool;
      DB_10_11_25 : Bool;
      DB_10_11_26 : Bool;
      DB_10_11_27 : Bool;
      DB_10_11_28 : Bool;
      DB_10_11_29 : Bool;
      DB_10_11_30 : Bool;
      DB_10_11_31 : Bool;
      DB_10_11_32 : Bool;
      DB_10_11_33 : Bool;
      DB_10_11_34 : Bool;
      DB_10_11_35 : Bool;
      DB_10_11_36 : Bool;
      DB_10_11_37 : Bool;
      DB_10_11_38 : Bool;
      DB_10_11_39 : Bool;
      DB_10_11_40 : Bool;
      DB_10_11_41 : Bool;
      DB_10_11_42 : Bool;
      DB_10_11_43 : Bool;
      DB_10_11_44 : Bool;
      DB_10_11_45 : Bool;
      DB_10_11_46 : Bool;
      DB_10_11_47 : Bool;
      DB_10_11_48 : Bool;
      DB_10_11_49 : Bool;
      DB_10_11_50 : Bool;
      DB_10_11_51 : Bool;
      DB_10_11_52 : Bool;
      DB_10_11_53 : Bool;
      DB_10_11_54 : Bool;
      DB_10_11_55 : Bool;
      DB_10_11_56 : Bool;
      DB_10_11_57 : Bool;
      DB_10_11_58 : Bool;
      DB_10_11_59 : Bool;
      DB_10_11_60 : Bool;
      DB_10_11_61 : Bool;
      DB_10_11_62 : Bool;
      DB_10_11_63 : Bool;
      DB_10_11_64 : Bool;
      DB_10_11_65 : Bool;
      DB_10_11_66 : Bool;
      DB_10_11_67 : Bool;
      DB_10_11_68 : Bool;
      DB_10_11_69 : Bool;
      DB_10_11_70 : Bool;
      DB_10_11_71 : Bool;
      DB_10_11_72 : Bool;
      DB_10_11_73 : Bool;
      DB_10_11_74 : Bool;
      DB_10_11_75 : Bool;
      DB_10_11_76 : Bool;
      DB_10_11_77 : Bool;
      DB_10_11_78 : Bool;
      DB_10_11_79 : Bool;
      DB_10_11_80 : Bool;
      DB_10_11_81 : Bool;
      DB_10_11_82 : Bool;
      DB_10_11_83 : Bool;
      DB_10_11_84 : Bool;
      DB_10_11_85 : Bool;
      DB_10_11_86 : Bool;
      DB_10_11_87 : Bool;
      DB_10_11_88 : Bool;
      DB_10_11_89 : Bool;
      DB_10_11_90 : Bool;
      DB_10_11_91 : Bool;
      DB_10_11_92 : Bool;
      DB_10_11_93 : Bool;
      DB_10_11_94 : Bool;
      DB_10_11_95 : Bool;
      DB_10_11_96 : Bool;
      DB_10_11_97 : Bool;
      DB_10_11_98 : Bool;
      DB_10_11_99 : Bool;
   END_VAR
BEGIN
END_DATA_BLOCK

DATA_BLOCK "FB11_DATA_ALARM_FB_DB"   // DB11
{ S7_Optimized_Access := 'FALSE' }
VERSION : 0.1
// stored: InstanceOfName FB11_DATA_ALARM_FB
"FB11_DATA_ALARM_FB"
BEGIN
END_DATA_BLOCK

DATA_BLOCK "HMI_OUT_BOOL"   // DB14
{ S7_Optimized_Access := 'FALSE' }